// TIA Portal project "XSFW_TIA60401_A2" (V13)

(* hardware
DEVICE "SIMATIC 300(1)"  S7-300 station
   slot 0: "UR"  Rail  6ES7 390-1***0-0AA0
   slot 2: "CPU 315-2PN/DP"  CPU 315-2 PN/DP  6ES7 315-2EH14-0AB0  V3.1
      slot 2: "PN-IO"  PN-IO
         slot 1: "Puerto 1"  Port
         slot 2: "Puerto 2"  Port
   slot 4: "DI32xDC24V"  DI32xDC24V  6ES7 321-1BL00-0AA0
   slot 5: "DI32xDC24V_1"  DI32xDC24V  6ES7 321-1BL00-0AA0
   slot 6: "DI32xDC24V_2"  DI32xDC24V  6ES7 321-1BL00-0AA0
   slot 7: "DO32xDC24V/0.5A"  DO32xDC24V/0.5A  6ES7 322-1BL00-0AA0
   slot 8: "DO32xDC24V/0.5A_1"  DO32xDC24V/0.5A  6ES7 322-1BL00-0AA0
   slot 9: "AI8x13Bit"  AI8x13Bit  6ES7 331-1KF02-0AB0
   slot 10: "AI8x13Bit_1"  AI8x13Bit  6ES7 331-1KF02-0AB0
DEVICE "HMI-Chillers"  TP900 Comfort
   slot 0: "HMI"  HMI  6AV2 124-0JC01-0AX0  11.0.0
   slot 1: "HMI_RT_3"  TP900 Comfort  6AV2 124-0JC01-0AX0  11.0.0
   slot 5: "IE_CP_1"  PROFINET interface  IE_CP  V7.1.0
      slot 1: "PROFINET_Interfaz_1"  HMI IE SUBMODULE
         slot 1: "PORT_1"  HMI IE PORTMODULE 1  1.0.0.0
         slot 2: "PORT_2"  HMI IE PORTMODULE 1  1.0.0.0
   slot 7: "MPI/DP_CP_1"  HMI MPIDP  MPI-DP_CP  1.0.0.0
DEVICE "IM153-4PN"  S7-300 station
   slot 0: "UR"  Rail  6ES7 390-1***0-0AA0
   slot 0: "IM153-4PN"  IM 153-4PN  6ES7 153-4AA01-0XB0  V2.0
   slot 1: "DI32xDC24V"  DI32xDC24V  6ES7 321-1BL00-0AA0
   slot 2: "DI32xDC24V_2"  DI32xDC24V  6ES7 321-1BL00-0AA0
   slot 3: "DI32xDC24V_3"  DI32xDC24V  6ES7 321-1BL00-0AA0
   slot 4: "DO32xDC24V/0.5A_2"  DO32xDC24V/0.5A  6ES7 322-1BL00-0AA0
   slot 5: "DO32xDC24V/0.5A"  DO32xDC24V/0.5A  6ES7 322-1BL00-0AA0
   slot 6: "AI8x12Bit"  AI8 x 12 bits  6ES7 331-7KF02-0AB0
DEVICE "Cavaleto"  TP1200 Comfort
   slot 0: "HMI"  HMI  6AV2 124-0MC01-0AX0  13.0.1.0
   slot 1: "HMI_RT_1"  TP1200 Comfort  6AV2 124-0MC01-0AX0  13.0.1.0
   slot 5: "Cavaleto.IE_CP_1"  Interfaz PROFINET
      slot 1: "Interfaz PROFINET_1"  Interfaz PROFINET
         slot 1: "Port_1"  Port
         slot 2: "Port_2"  Port
   slot 7: "Cavaleto.MPI/DP_CP_1"  Interfaz MPI/DP
*)

// ===== PLC "CPU 315-2PN/DP"  CPU 315-2 PN/DP =====
// protected blocks, not shown: "FB_CTR_MOT", "FB_PRC_ALA", "FC_ANIM_MOTOR", "FC_CH_AI", "FC_MAQ_EST_16", "FC_PRC_ALA2", "FC_PRC_ALA3"

VAR_GLOBAL   // PLC tag table "Tabla de variables estándar"
   "Tag_1" AT %M7.0 : Bool;
   "Tag_2" AT %M7.1 : Bool;
   "Tag_3" AT %M7.2 : Bool;
   "Tag_4" AT %M7.3 : Bool;
   "Tag_5" AT %M7.4 : Bool;
   "Tag_6" AT %M500.0 : Bool;
   "Tag_7" AT %M900.0 : Bool;
   "Tag_9" AT %T15 : Timer;
   "Tag_10" AT %T16 : Timer;
   "Tag_11" AT %M55.0 : Bool;
   "Tag_12" AT %M330.3 : Bool;
   "Tag_13" AT %T80 : Timer;
   "flReqMch2" AT %M70.1 : Bool;
   "flReqMch3" AT %M70.2 : Bool;
   "flReqMch4" AT %M70.3 : Bool;
   "flReqMch5" AT %M70.4 : Bool;
   "Tag_18" AT %T62 : Timer;
   "Tag_19" AT %T61 : Timer;
   "Tag_20" AT %T60 : Timer;
   "Tag_21" AT %T70 : Timer;
   "Tag_22" AT %T71 : Timer;
   "Tag_23" AT %T72 : Timer;
   "Tag_24" AT %T73 : Timer;
   "Tag_25" AT %T74 : Timer;
   "Tag_26" AT %T24 : Timer;
   "Tag_27" AT %T10 : Timer;
   "Tag_28" AT %T11 : Timer;
   "Tag_29" AT %T12 : Timer;
   "Tag_30" AT %T13 : Timer;
   "Tag_31" AT %T14 : Timer;
   "Tag_32" AT %T26 : Timer;
   "Tag_33" AT %T28 : Timer;
   "Tag_34" AT %T30 : Timer;
   "Tag_35" AT %T32 : Timer;
   "Tag_36" AT %T34 : Timer;
   "Tag_37" AT %Q100.5 : Bool;
   "Tag_38" AT %M0.4 : Bool;
   "Tag_39" AT %Q104.4 : Bool;
   "Tag_40" AT %Q104.5 : Bool;
   "Tag_41" AT %Q101.1 : Bool;
   "Tag_42" AT %Q101.2 : Bool;
   "Tag_43" AT %Q101.3 : Bool;
   "Tag_44" AT %Q101.4 : Bool;
   "Tag_45" AT %Q101.5 : Bool;
   "Tag_46" AT %Q101.6 : Bool;
   "Tag_47" AT %Q101.7 : Bool;
   "Tag_48" AT %M25.0 : Bool;
   "Tag_49" AT %M25.1 : Bool;
   "Tag_50" AT %M25.2 : Bool;
   "Tag_51" AT %T35 : Timer;
   "Tag_52" AT %Q102.3 : Bool;
   "Tag_53" AT %Q102.4 : Bool;
   "Tag_54" AT %Q102.5 : Bool;
   "Tag_103" AT %M0.7 : Bool;
   "Tag_115" AT %M0.2 : Bool;
   "Tag_146" AT %M0.6 : Bool;
   "Tag_154" AT %M50.0 : Bool;
   "Tag_155" AT %M2.1 : Bool;
   "Tag_156" AT %M50.3 : Bool;
   "Tag_157" AT %M2.2 : Bool;
   "Tag_158" AT %M50.5 : Bool;
   "Tag_159" AT %M2.0 : Bool;
   "Tag_160" AT %Q69.1 : Bool;   // -
   "Tag_161" AT %M55.7 : Bool;
   "Tag_162" AT %M55.6 : Bool;
   "Latch_FT1" AT %M80.0 : Bool;   // Retención Flanco en Flujostato
   "Permiso_NO_FT1" AT %M80.1 : Bool;   // Permiso para trabajar sin FT1
   "Auxiliar_FT1" AT %M80.2 : Bool;
   "Auxiliar_Timer_FT1" AT %M80.3 : Bool;
   "Aviso 1" AT %M82.0 : Bool;
   "Aviso 2" AT %M82.1 : Bool;
   "Aviso 3" AT %M82.2 : Bool;
   "Aviso 4" AT %M82.3 : Bool;
   "Aviso 5" AT %M82.4 : Bool;
   "Aviso 13" AT %M82.6 : Bool;
   "Aviso 14" AT %M82.7 : Bool;
   "Aviso 23" AT %M83.0 : Bool;
   "Aviso 24" AT %M83.1 : Bool;
   "Aviso25" AT %M83.2 : Bool;
   "Aviso 26" AT %M83.3 : Bool;
   "Aviso 27" AT %M83.4 : Bool;
   "UltimoCmdMarcha" AT %M90.0 : Bool;
   "Tag_163" AT %T87 : Timer;
   "NotFirstScan" AT %M900.1 : Bool;
   "Tag_14" AT %M760.1 : Bool;
   "Tag_15" AT %M760.2 : Bool;
   "EnclavCompAltaConFlujostato" AT %M93.4 : Bool;
   "EstadoMantMC001" AT %MB761 : Byte;
   "EstadoMantMC002" AT %MB762 : Byte;
   "EstadoMantMC003" AT %MB763 : Byte;
   "EstadoMantMC004" AT %MB764 : Byte;
   "EstadoMantMC005" AT %MB765 : Byte;
   "EstadoMantMC006" AT %MB766 : Byte;
   "LimiteMantMC001_1" AT %M761.0 : Bool;
   "LimiteMantMC001_2" AT %M761.1 : Bool;
   "LimiteMantMC002_1" AT %M762.0 : Bool;
   "LimiteMantMC002_2" AT %M762.1 : Bool;
   "LimiteMantMC003_1" AT %M763.0 : Bool;
   "LimiteMantMC003_2" AT %M763.1 : Bool;
   "LimiteMantMC004_1" AT %M764.0 : Bool;
   "LimiteMantMC004_2" AT %M764.1 : Bool;
   "LimiteMantMC005_1" AT %M765.0 : Bool;
   "LimiteMantMC005_2" AT %M765.1 : Bool;
   "LimiteMantMC006_1" AT %M766.0 : Bool;
   "LimiteMantMC006_2" AT %M766.1 : Bool;
   "ProxMantMC001_1" AT %MD768 : DInt;
   "ProxMantMC002_1" AT %MD772 : DInt;
   "ProxMantMC003_1" AT %MD776 : DInt;
   "ProxMantMC004_1" AT %MD780 : DInt;
   "ProxMantMC005_1" AT %MD784 : DInt;
   "ProxMantMC006_1" AT %MD788 : DInt;
   "ProxMantMC001_2" AT %MD792 : DInt;
   "ProxMantMC002_2" AT %MD796 : DInt;
   "ProxMantMC003_2" AT %MD800 : DInt;
   "ProxMantMC004_2" AT %MD804 : DInt;
   "ProxMantMC005_2" AT %MD808 : DInt;
   "ProxMantMC006_2" AT %MD812 : DInt;
   "ProxMantMS050" AT %MD816 : DInt;
   "ProxMantMS051" AT %MD820 : DInt;
   "ProxMantMS052" AT %MD824 : DInt;
   "ProxMantMS053" AT %MD828 : DInt;
   "LimiteMantMS050" AT %M767.0 : Bool;
   "LimiteMantMS051" AT %M767.1 : Bool;
   "LimiteMantMS052" AT %M767.2 : Bool;
   "LimiteMantMS053" AT %M767.3 : Bool;
   "LimiteMantMS054_1" AT %M832.0 : Bool;
   "LimiteMantMS055_1" AT %M832.2 : Bool;
   "LimiteMantMS056_1" AT %M832.4 : Bool;
   "LimiteMantMS054_2" AT %M832.1 : Bool;
   "LimiteMantMS055_2" AT %M832.3 : Bool;
   "LimiteMantMS056_2" AT %M832.5 : Bool;
   "ProxMantMC060_1" AT %MD834 : DInt;
   "ProxMantMC061_1" AT %MD838 : DInt;
   "ProxMantMC062_1" AT %MD842 : DInt;
   "ProxMantMC063_1" AT %MD846 : DInt;
   "ProxMantMC064_1" AT %MD850 : DInt;
   "ProxMantMC065_1" AT %MD854 : DInt;
   "ProxMantMC060_2" AT %MD858 : DInt;
   "ProxMantMC061_2" AT %MD862 : DInt;
   "ProxMantMC062_2" AT %MD866 : DInt;
   "ProxMantMC063_2" AT %MD870 : DInt;
   "ProxMantMC064_2" AT %MD874 : DInt;
   "ProxMantMC065_2" AT %MD878 : DInt;
   "ProxMantMC060_3" AT %MD882 : DInt;
   "ProxMantMC061_3" AT %MD886 : DInt;
   "ProxMantMC062_3" AT %MD890 : DInt;
   "ProxMantMC063_3" AT %MD894 : DInt;
   "ProxMantMC064_3" AT %MD910 : DInt;
   "ProxMantMC065_3" AT %MD914 : DInt;
   "ProxMantMC060_4" AT %MD918 : DInt;
   "ProxMantMC061_4" AT %MD922 : DInt;
   "ProxMantMC062_4" AT %MD926 : DInt;
   "ProxMantMC063_4" AT %MD930 : DInt;
   "ProxMantMC064_4" AT %MD934 : DInt;
   "ProxMantMC065_4" AT %MD938 : DInt;
   "ProxMantMC060_5" AT %MD942 : DInt;
   "ProxMantMC061_5" AT %MD946 : DInt;
   "ProxMantMC062_5" AT %MD950 : DInt;
   "ProxMantMC063_5" AT %MD954 : DInt;
   "ProxMantMC064_5" AT %MD958 : DInt;
   "ProxMantMC065_5" AT %MD962 : DInt;
   "LimiteMantMC060_1" AT %M901.0 : Bool;
   "LimiteMantMC060_2" AT %M901.1 : Bool;
   "LimiteMantMC060_3" AT %M901.2 : Bool;
   "LimiteMantMC060_4" AT %M901.3 : Bool;
   "LimiteMantMC060_5" AT %M901.4 : Bool;
   "LimiteMantMC061_1" AT %M902.0 : Bool;
   "LimiteMantMC061_2" AT %M902.1 : Bool;
   "LimiteMantMC061_3" AT %M902.2 : Bool;
   "LimiteMantMC061_4" AT %M902.3 : Bool;
   "LimiteMantMC061_5" AT %M902.4 : Bool;
   "LimiteMantMC062_1" AT %M903.0 : Bool;
   "LimiteMantMC062_2" AT %M903.1 : Bool;
   "LimiteMantMC062_3" AT %M903.2 : Bool;
   "LimiteMantMC062_4" AT %M903.3 : Bool;
   "LimiteMantMC062_5" AT %M903.4 : Bool;
   "LimiteMantMC063_1" AT %M904.0 : Bool;
   "LimiteMantMC063_2" AT %M904.1 : Bool;
   "LimiteMantMC063_3" AT %M904.2 : Bool;
   "LimiteMantMC063_4" AT %M904.3 : Bool;
   "LimiteMantMC063_5" AT %M904.4 : Bool;
   "LimiteMantMC064_1" AT %M905.0 : Bool;
   "LimiteMantMC064_2" AT %M905.1 : Bool;
   "LimiteMantMC064_3" AT %M905.2 : Bool;
   "LimiteMantMC064_4" AT %M905.3 : Bool;
   "LimiteMantMC064_5" AT %M905.4 : Bool;
   "LimiteMantMC065_1" AT %M906.0 : Bool;
   "LimiteMantMC065_2" AT %M906.1 : Bool;
   "LimiteMantMC065_3" AT %M906.2 : Bool;
   "LimiteMantMC065_4" AT %M906.3 : Bool;
   "LimiteMantMC065_5" AT %M906.4 : Bool;
   "EstadoMantMC060" AT %MB901 : Byte;
   "EstadoMantMC061" AT %MB902 : Byte;
   "EstadoMantMC062" AT %MB903 : Byte;
   "EstadoMantMC063" AT %MB904 : Byte;
   "EstadoMantMC064" AT %MB905 : Byte;
   "ProxMantMS054_1" AT %MD966 : DInt;
   "ProxMantMS054_2" AT %MD970 : DInt;
   "ProxMantMS055_1" AT %MD974 : DInt;
   "ProxMantMS055_2" AT %MD978 : DInt;
   "EstadoMantSecBaja" AT %MB832 : Byte;
   "EnclavCompAltaPorTemp" AT %M93.5 : Bool;
   "FallTempCritEnclav" AT %M93.6 : Bool;
   "EntAnalCaudal" AT %IW266 : Word;
   "Tag_57" AT %MW982 : Word;
   "Tag_59" AT %MW984 : Word;
   "Tag_8" AT %M982.0 : Bool;
   "Tag_16" AT %M982.1 : Bool;
   "EntAnalPotencia" AT %IW264 : Word;
   "Tag_17" AT %T90 : Timer;
   "Tag_55" AT %T91 : Timer;
   "Tag_56" AT %M100.0 : Bool;
   "Tag_58" AT %M1000.0 : Bool;
   "Tag_60" AT %MW1010 : S5Time;
   "Tag_61" AT %MW1012 : S5Time;
   "MC003_EVP" AT %Q7.2 : Bool;   // Purga Bellis
   "Tag_63" AT %M1000.1 : Bool;
   "Tag_64" AT %T92 : Timer;
   "Tag_65" AT %T93 : Timer;
   "Tag_66" AT %MW1014 : S5Time;
   "Tag_67" AT %MW1016 : S5Time;
   "MC001_EVP" AT %Q7.3 : Bool;   // Purga ABC2
   "Tag_69" AT %M1000.2 : Bool;
   "Tag_70" AT %T94 : Timer;
   "Tag_71" AT %T95 : Timer;
   "Tag_72" AT %MW1018 : S5Time;
   "Tag_73" AT %MW1020 : S5Time;
   "MC002_EVP" AT %Q7.4 : Bool;   // Purga ABC3
   "Tag_75" AT %T96 : Timer;
   "Tag_76" AT %T97 : Timer;
   "MC004_EVP" AT %Q7.5 : Bool;   // Purga ABC4
   "Tag_78" AT %T98 : Timer;
   "Tag_79" AT %T99 : Timer;
   "MC005_EVP" AT %Q7.6 : Bool;   // Purga ABC5
   "Tag_62" AT %T100 : Timer;
   "MC006_EVP" AT %Q7.7 : Bool;   // Purga ABC1
   "Tag_68" AT %M1000.7 : Bool;
   "Tag_74" AT %T101 : Timer;
   "Tag_77" AT %T102 : Timer;
   "Tag_80" AT %T103 : Timer;
   "Tag_81" AT %T104 : Timer;
   "Tag_82" AT %T105 : Timer;
   "Tag_83" AT %T106 : Timer;
   "Tag_84" AT %T107 : Timer;
   "Tag_85" AT %I78.1 : Bool;
END_VAR

VAR_GLOBAL   // PLC tag table "STEP7 classic symbols"
   "MS055_MANT" AT %A4.1 : Bool;   // S BAJA SULLAIR 2-SEÑAL MODO MANTENIMIENTO / Secador 6 - SRD 1000 - Salida de Mantenimiento
   "MS055_Marcha" AT %A4.7 : Bool;   // S BAJA SULLAIR 2-CONTACTOR / Secador 6 - SRD 1000 - Salida de Marcha
   "MC006_TTB" AT %E2.2 : Bool;   // M COMPRESOR ALTA ABC1-TERMOSTATO AGUA / Secador 7 falla termico
   "MC006_TTA" AT %E2.3 : Bool;   // M COMPRESOR ALTA ABC1-TERMOSTATO AIRE / secador 8 falla termico
   "MT007-CO" AT %E66.0 : Bool;   // B SOPLADO L1-CONFIRMACIÓN DE MARCHA / Bomba Principal Chiller Soplado - Confirmación de Marcha
   "MT007-Marcha" AT %A66.0 : Bool;   // B SOPLADO L1-CONTACTOR / Accionamiento Bomba Intercambiador LINEA 1
   "MT007-TO" AT %E66.1 : Bool;   // B SOPLADO L1-TÉRMICO / Bomba Principal Chiller Soplado - Falla de Térmico
   "MT008-CO" AT %E66.2 : Bool;   // B SOPLADO L3 & MANOMEC-CONFIRMACIÓN DE MARCHA / Bomba Backup Chiller Soplado - Confirmación de Marcha
   "MT008-Marcha" AT %A66.1 : Bool;   // B SOPLADO L3 & MANOMEC-CONTACTOR / Accionamiento Bomba Intercambiador LINEA 2 Y MANOMEC
   "MT008-TO" AT %E66.3 : Bool;   // B SOPLADO L3 & MANOMEC-TÉRMICO / Bomba Backup Chiller Soplado - Falla de Térmico
   "MT009-CO" AT %E66.4 : Bool;   // B INT L3 Y L5-CONFIRMACIÓN DE MARCHA / Bomba Principal Chiller Envasado - Confirmación de Marcha
   "MT009-Marcha" AT %A66.2 : Bool;   // B INT L3 Y L5-CONTACTOR / Accionamiento Bomba Intercambiador LINEA 3 Y LINEA 5
   "MS052-TO" AT %E1.6 : Bool;   // M SECADOR ALTA ABC2-TÉRMICO / Secador 3-ABC 3- falla termico
   "MS052-VS1" AT %E9.4 : Bool;   // M SECADOR ALTA ABC2-PULSADOR PARADA / Secador 3 -ABC 3 - Falla de seguridades
   "MS052_MANT" AT %A3.6 : Bool;   // M SECADOR ALTA ABC2-SEÑAL MODO MANTENIMIENTO / Secador 2 - ABC 2 - Salida de Mantenimiento
   "FlancoMan2" AT %M322.7 : Bool;
   "FlancoMan3" AT %M323.0 : Bool;
   "FlancoMan4" AT %M323.1 : Bool;
   "FlancoMan5" AT %M323.2 : Bool;
   "FlancoManP1" AT %M323.3 : Bool;
   "FlancoManP2" AT %M323.4 : Bool;
   "FlancoManP3" AT %M323.5 : Bool;
   "FlancoManP4" AT %M323.6 : Bool;
   "FlancoManP5" AT %M323.7 : Bool;
   "TLUZ" AT %T17 : Timer;   // Tiempo Iluminación encendida
   "TOFF_SP1" AT %T44 : Timer;   // TOFF sopladora 1
   "TOFF_SP2" AT %T45 : Timer;   // TOFF Sopladora 2
   "TOFF_SP3" AT %T46 : Timer;   // TOFF Sopladora 3
   "TRetVCmp1" AT %T51 : Timer;   // Timer Retardo arranque de valvulas Compresor 1
   "TRetVCmp2" AT %T47 : Timer;   // Timer Retardo arranque de valvulas Compresor 2
   "TRetVCmp3" AT %T48 : Timer;   // Timer Retardo arranque de valvulas Compresor 3
   "TRetVCmp4" AT %T49 : Timer;   // Timer Retardo arranque de valvulas Compresor 4
   "TV1" AT %T53 : Timer;   // Timeout estando en vacío 1
   "TV2" AT %T36 : Timer;   // Timeout estando en vacío 2
   "TV3" AT %T37 : Timer;   // Timeout estando en vacío 3
   "TV4" AT %T38 : Timer;   // Timeout estando en vacío 4
   "FlaAux3" AT %M300.2 : Bool;   // Auxiliar arranque MC003
   "FlaAux4" AT %M300.3 : Bool;   // Auxiliar arranque MC004
   "FlaAux5" AT %M300.4 : Bool;   // Auxiliar arranque MC005
   "FlaAuxB1" AT %M300.5 : Bool;   // Auxiliar arranque MC061
   "FlaAuxB2" AT %M300.6 : Bool;   // Auxiliar arranque MC062
   "FlaAuxB3" AT %M300.7 : Bool;   // Auxiliar arranque MC063
   "FlaAuxB4" AT %M301.0 : Bool;   // Auxiliar arranque MC064
   "FlancoAuto1" AT %M324.0 : Bool;
   "FlancoAuto2" AT %M324.1 : Bool;
   "MP011-CO" AT %E67.2 : Bool;   // B BACKUP CH. SOPLADO-CONFIRMACIÓN DE MARCHA / Bomba Intercambiador LINEA 2 Y MANOMEC - Confirmación de Marcha
   "MP011-Marcha" AT %A66.5 : Bool;   // B BACKUP CH. SOPLADO-CONTACTOR / Accionamiento Bomba Backup Chiller Soplado
   "MP011-TO" AT %E67.3 : Bool;   // B BACKUP CH. SOPLADO-TÉRMICO / Bomba Intercambiador LINEA 2 Y MANOMEC - Falla de Térmico
   "MP012-CO" AT %E67.4 : Bool;   // B PRINC CH. ENVASADO-CONFIRMACIÓN DE MARCHA / Bomba Intercambiador LINEA 3 Y LINEA 5 - Confirmación de Marcha
   "MP012-Marcha" AT %A66.6 : Bool;   // B PRINC CH. ENVASADO-CONTACTOR / Accionamiento Bomba Principal Chiller Envasado
   "ArrMC061" AT %T81 : Timer;   // Timer arranque MC061
   "ArrMC062" AT %T82 : Timer;   // Timer arranque MC062
   "ArrMC063" AT %T83 : Timer;   // Timer arranque MC063
   "ArrMC064" AT %T84 : Timer;   // Timer arranque MC064
   "Arracando_MC002" AT %T27 : Timer;
   "Arrancando_MC001" AT %T25 : Timer;   // Delay para meter EV
   "Arrancando_MC004" AT %T31 : Timer;
   "Arrancando_MC005" AT %T33 : Timer;
   "Arrancando_mc003" AT %T29 : Timer;
   "BBA POZO" AT %A0.4 : Bool;   // BOMBA POZO- / BOMBA DE POZO
   "BMBTON2" AT %M69.3 : Bool;   // Bomba de torre 2 en funcionamiento
   "BMBTON2BMBTON" AT %M69.2 : Bool;   // Bomba de torre en funcionamiento
   "MC061-TO" AT %E11.5 : Bool;   // M COMPR BAJA SULLAIR 1-TÉRMICO / Compresor Baja SULL 1 - Falla de termico
   "MC005_ConfPurga" AT %E11.6 : Bool;   // ABC5 - Confirmación de electroválvula de purga. / Compresor Baja SULL 1 - Falla de seguridades
   "MC061_MANT" AT %A1.4 : Bool;   // M COMPR BAJA SULLAIR 1-SEÑAL MODO MANTENIMIENTO / Compresor Sullair1 Salida mantenimiento
   "MC061_MARCHA" AT %A1.5 : Bool;   // M COMPR BAJA SULLAIR 1-CONTACTOR / Comrpesor Sullair1 Salida de marcha
   "MC062-CO" AT %E10.3 : Bool;   // M COMPR BAJA SULLAIR 0-CONFIRMACIÓN DE MARCHA / Compresor Baja SULL 0- Conf. Marcha
   "MC062-TO" AT %E10.4 : Bool;   // M COMPR BAJA SULLAIR 0-TÉRMICO / Compresor Baja SULL 0- Falla de termico
   "MC062-VS1" AT %E10.5 : Bool;   // M COMPR BAJA SULLAIR 0-PULSADOR PARADA / Compresor Baja SULL 0- Falla de Seguridades
   "MC062_MANT" AT %A1.6 : Bool;   // M COMPR BAJA SULLAIR 0-SEÑAL MODO MANTENIMIENTO / Compresor XXX salida de mantenimiento
   "MC062_MARCHA" AT %A1.7 : Bool;   // M COMPR BAJA SULLAIR 0-CONTACTOR / Compresor XXX salida de marcha EX61
   "MC063-CO" AT %E10.6 : Bool;   // M COMPR BAJA ATLAS 3-CONFIRMACIÓN DE MARCHA / Compresor Baja ATLAS 3 - Conf.Marcha
   "MC063-TO" AT %E10.7 : Bool;   // M COMPR BAJA ATLAS 3-TÉRMICO / Compresor Baja ATLAS 3 - Falla de termico
   "IndicadorCmpAlta" AT %M310.4 : Bool;   // Indicador Aviso en Compresores de alta
   "IndicadorCmpBaja" AT %M310.2 : Bool;   // Indicador Aviso en Compresores de baja
   "IndicadorSecAlta" AT %M310.5 : Bool;   // Indicador Aviso en Secadores de alta
   "IndicadorSecBaja" AT %M310.3 : Bool;   // Indicador Aviso en Secadores de baja
   "IndicadorTorresCav" AT %M310.6 : Bool;   // Indicador Aviso en Torres cavalleto
   "IndicadorTorresCh" AT %M310.1 : Bool;   // Indicador Aviso en torres chillers
   "MC001" AT %A0.6 : Bool;   // M COMPRESOR ALTA ABC2-CONTACTOR / Compresor ABC2- Marcha-
   "MC001-CO" AT %E2.5 : Bool;   // M COMPRESOR ALTA ABC2-CONFIRMACIÓN DE MARCHA / Compresor ABC2-Confirmacion Marcha-
   "MC001-TO" AT %E2.6 : Bool;   // M COMPRESOR ALTA ABC2-TÉRMICO / Compresor ABC2-Falla Termico-
   "MC001_EV" AT %A2.0 : Bool;   // M COMPRESOR ALTA ABC2-ELECTROVÁLVULA / Electrovalvula libera carga MC001 (ABC2)
   "MC001_MANT" AT %A2.5 : Bool;   // M COMPRESOR ALTA ABC2-SEÑAL MODO MANTENIMIENTO / Compresor MC001 Salida Mantenimiento
   "MC002_ConfPurga" AT %E1.1 : Bool;   // ABC3 - Confirmación de electroválvula de purga. / Bomba de pozo -falla termico-
   "flReqMch1" AT %M70.0 : Bool;   // Flanco requerimiento de marcha compresor 1
   "TRetVCmp5" AT %T50 : Timer;   // Timer Retardo arranque de valvulas Compresor 5
   "FlancoTSinReq4" AT %M325.6 : Bool;
   "FlancoTSinReq5" AT %M325.7 : Bool;
   "FallaSensorTorresCH" AT %M77.7 : Bool;   // Falla en Sensor de Temperatura Torres de Chillers
   "FlaAux1" AT %M300.0 : Bool;   // Auxiliar arranque MC001
   "FlaAux2" AT %M300.1 : Bool;   // Auxiliar arranque MC002
   "Parada-MC062" AT %A6.0 : Bool;   // M COMPR BAJA SULLAIR 0-ORDEN PARADA / Parada MC062
   "Parada-MC063" AT %A5.7 : Bool;   // M COMPR BAJA ATLAS 3-ORDEN PARADA / Parada MC063
   "Parada-MC064" AT %A5.6 : Bool;   // M COMPR BAJA ATLAS 2-ORDEN PARADA / Parada MC064
   "P_PresALTA" AT %EW254 : Word;   // PresiónALTA
   "P_PresAlta2" AT %EW258 : Word;   // PresiónAlta2
   "P_PresBaja" AT %EW260 : Word;   // Presión Baja
   "Puls.Iluminati" AT %E7.5 : Bool;   // ILUMINACION-PULSADOR / Pulsador Iluminacion
   "Pulso0,5_Seg" AT %M1.0 : Bool;
   "Pulso100_Mseg" AT %M0.3 : Bool;
   "Pulso10_Seg" AT %M1.3 : Bool;
   "Pulso1_Seg" AT %M1.1 : Bool;
   "ErrCMQ1" AT %M320.5 : Bool;   // Error Concatenadoras Compresor 1
   "ErrCMQ2" AT %M320.6 : Bool;   // Error Concatenadoras Compresor 2
   "ErrCMQ3" AT %M320.7 : Bool;   // Error Concatenadoras Compresor 3
   "ErrCMQ4" AT %M321.0 : Bool;   // Error Concatenadoras Compresor 4
   "ErrCMQ5" AT %M321.1 : Bool;   // Error Concatenadoras Compresor 5
   "ErrCMQG" AT %M321.3 : Bool;   // Error Concatenadoras General
   "ErrPMQ1" AT %M320.0 : Bool;   // Error Prioritarias Compresor 1
   "ErrPMQ2" AT %M320.1 : Bool;   // Error Prioritarias Compresor 2
   "ErrPMQ3" AT %M320.2 : Bool;   // Error Prioritarias Compresor 3
   "ErrPMQ4" AT %M320.3 : Bool;   // Error Prioritarias Compresor 4
   "ErrPMQ5" AT %M320.4 : Bool;   // Error Prioritarias Compresor 5
   "BoosterAnimaMotor" AT %MB11 : Byte;   // Byte Animación Motor Booster
   "BoostMoManten" AT %M10.0 : Bool;   // Booster en modo Mantenimiento
   "BoostMoManual" AT %M10.1 : Bool;   // Booster en modo Manual
   "BoostMoAutoma" AT %M10.2 : Bool;   // Booster en modo Automático
   "BoosterAlarma" AT %M10.3 : Bool;   // Booster con Alarma Memorizada
   "BoostOrdMarch" AT %M10.4 : Bool;   // Booster con Orden de Marcha
   "BoostPlsManten" AT %M10.5 : Bool;   // Booster Pulsa Mantenimiento desde HMI
   "iConfMarBooster" AT %E3.7 : Bool;   // M BOOSTER 1-CONFIRMACIÓN DE MARCHA / Confirmaciónes Marcha serie motores Booster
   "iGMBooster" AT %E4.0 : Bool;   // M BOOSTER 1-GUARDAMOTOR / Confirmaciónes Guardamotores serie motores Booster
   "iPresostCtrl" AT %E7.6 : Bool;   // BOOSTERS (LOS DOS)-PRESOSTATO / Presostato de Control para Booster
   "iPresostPA" AT %E7.7 : Bool;   // BOOSTERS (LOS DOS)-PRESOSTATO PRESION ALTA / Presostato de "Presión Alta" para Booster
   "oMarBooster" AT %A7.0 : Bool;   // BOOSTER-CONTACTOR / Accionamiento Contactor Booster
   "FiltroPCtrlBooster" AT %T18 : Timer;   // Filtro de Presión de Control de Booster
   "FiltroPABooster" AT %T19 : Timer;   // Filtro de Presión Alta de Booster
   "Boost2OrdMarch" AT %M12.5 : Bool;   // Booster 2 con Orden de Marcha
   "Booster2Alarma" AT %M12.4 : Bool;   // Booster 2 con Alarma Memorizada
   "Boost2MoAutoma" AT %M12.3 : Bool;   // Booster 2 en modo Automático
   "Boost2MoManual" AT %M12.2 : Bool;   // Booster 2 en modo Manual
   "Boost2MoManten" AT %M12.1 : Bool;   // Booster 2 en modo Mantenimiento
   "BoostHabilit" AT %M12.0 : Bool;   // Habilitación Booster desde HMI
   "Boost2PlsManual" AT %M12.7 : Bool;   // Booster 2 Pulsa Manual desde HMI
   "Boost2PlsManten" AT %M12.6 : Bool;   // Booster 2 Pulsa Mantenimiento desde HMI
   "ReservaBooster_5" AT %M13.6 : Bool;
   "ReservaBooster_4" AT %M13.5 : Bool;
   "ReservaBooster_3" AT %M13.4 : Bool;
   "MS052_Marcha" AT %A4.4 : Bool;   // M SECADOR ALTA ABC2-CONTACTOR / Secador 3 - ABC 3 - Salida de Marcha
   "MS053-CO" AT %E4.4 : Bool;   // M SECADOR ALTA FARGON-CONFIRMACIÓN DE MARCHA / Secador 4 - Fargon -Conf.Marcha
   "MS053-TO" AT %E1.7 : Bool;   // M SECADOR ALTA FARGON-TÉRMICO / Secador 4-FARGON -falla termico
   "MS053-VS1" AT %E9.5 : Bool;   // M SECADOR ALTA FARGON-PULSADOR PARADA / Secador 4 -ABC Grande - Falla de seguridades
   "MS053_MANT" AT %A3.7 : Bool;   // M SECADOR ALTA FARGON-SEÑAL MODO MANTENIMIENTO / Secador 4- FARGON- Salida de Mantenimiento
   "MS053_Marcha" AT %A4.5 : Bool;   // M SECADOR ALTA FARGON-CONTACTOR / Secador 4 - FARGON - Salida de marcha
   "MS054-CO" AT %E4.5 : Bool;   // S BAJA SULLAIR 1-CONFIRMACIÓN DE MARCHA / Secador 5 -SRD850 - Conf.Marcha
   "MC006-CO" AT %E2.0 : Bool;   // M COMPRESOR ALTA ABC1-CONFIRMACIÓN DE MARCHA / Secador 5 - SRD 850 -falla termico
   "iConfMarBooster2" AT %E9.6 : Bool;   // M BOOSTER 2-CONFIRMACIÓN DE MARCHA / Confirmación de marcha Booster 2
   "MS054_MANT" AT %A4.0 : Bool;   // S BAJA SULLAIR 1-SEÑAL MODO MANTENIMIENTO / Secador 5 - SRD850 - Salida de Mantenimiento
   "MS054_Marcha" AT %A4.6 : Bool;   // S BAJA SULLAIR 1-CONTACTOR / Secador 5 - SRD850 - Salida de Marcha
   "MS055-CO" AT %E4.6 : Bool;   // S BAJA SULLAIR 2-CONFIRMACIÓN DE MARCHA / Secador 6 - SRD1000 - Conf.Marcha
   "MC006_PTB" AT %E2.1 : Bool;   // M COMPRESOR ALTA ABC1-PRESOSTATO AGUA / Secador 6 - SRD 1000-falla termico
   "Corneta" AT %A3.3 : Bool;   // -ALARMA / Bubuzella
   "MP019-CO" AT %E68.2 : Bool;   // BOMBA 2-CONFIRMACIÓN DE MARCHA / Bomba 2 Torres Enfriamiento - Confirmación de Marcha
   "MP019-Marcha" AT %A67.1 : Bool;   // BOMBA 2-CONTACTOR / Accionamiento Bomba 2 Torres Enfriamiento
   "MP019-TO" AT %E68.3 : Bool;   // BOMBA 2-TÉRMICO / Bomba 2 Torres Enfriamiento - Falla de Térmico
   "MP019_PA" AT %E8.3 : Bool;   // BOMBA 2-PULSADOR MARCHA / Bomba 2 Torre Cavalleto Pulsador Arranque
   "MP019_PP" AT %E8.4 : Bool;   // BOMBA 2-PULSADOR PARADA / Bomba 2 Torre Cavalleto Pulsador Parada
   "FlancoNoFal2" AT %M324.6 : Bool;
   "FlancoNoFal3" AT %M324.7 : Bool;
   "FlancoNoFal4" AT %M325.0 : Bool;
   "FlancoNoFal5" AT %M325.1 : Bool;
   "FlancoOsc1s" AT %M326.0 : Bool;
   "FlancoPSop1" AT %M326.4 : Bool;
   "FlancoPSop2" AT %M326.5 : Bool;
   "FlancoPSop3" AT %M326.6 : Bool;
   "FlancoTSinReq1" AT %M325.3 : Bool;
   "FlancoTSinReq2" AT %M325.4 : Bool;
   "FlancoTSinReq3" AT %M325.5 : Bool;
   "TV5" AT %T39 : Timer;   // Timeout estando en vacío 5
   "TdesefMC060" AT %T54 : Timer;   // Tiempo desconexión efectiva MC060
   "TdesefMC061" AT %T55 : Timer;   // Tiempo desconexión efectiva MC061
   "TdesefMC062" AT %T56 : Timer;   // Tiempo desconexión efectiva MC062
   "TdesefMC063" AT %T57 : Timer;   // Tiempo desconexión efectiva MC063
   "TdesefMC064" AT %T58 : Timer;   // Tiempo desconexión efectiva MC064
   "P_TemCav" AT %EW256 : Word;   // Temperatura Torres Cavaleto
   "TempTorresCH" AT %MD52 : Real;   // Temperatura Torres de Chillers Escalada
   "P_TempTorresCHILL" AT %EW286 : Word;   // Temperatura de agua torres de enfriamiento chillers
   "MC006_PTA" AT %E2.4 : Bool;   // M COMPRESOR ALTA ABC1-PRESOSTATO ACEITE / tomascorrientes falla termico
   "Torre_PE" AT %E9.1 : Bool;   // TORRE ENFR-PULS PARADA EMER / Pulsador de emergencia torre de enfriamiento
   "FlancoDEC5" AT %M322.5 : Bool;
   "FlancoINC1" AT %M321.4 : Bool;
   "FlancoINC2" AT %M321.5 : Bool;
   "FlancoINC3" AT %M321.6 : Bool;
   "FlancoINC4" AT %M321.7 : Bool;
   "FlancoINC5" AT %M322.0 : Bool;
   "FlancoMan1" AT %M322.6 : Bool;
   "ReservaBooster_2" AT %M13.3 : Bool;
   "ReservaBooster_1" AT %M13.2 : Bool;
   "Boost2Habilit" AT %M13.1 : Bool;   // Habilitación Booster 2 desde HMI
   "Boost2PlsAutoma" AT %M13.0 : Bool;   // Booster 2 Pulsa Automático desde HMI
   "oMarBooster2" AT %A7.1 : Bool;   // BOOSTER 2-CONTACTOR / Accionamiento Contactor Booster 2
   "ReservaBooster_6" AT %M13.7 : Bool;
   "Booster2AnimaMotor" AT %MB14 : Byte;   // Byte Animación Motor Booster 2
   "PrioridadBoost2" AT %MW334 : Int;   // Prioridad de Arranque Booster 2
   "PrioridadBoost1" AT %MW332 : Int;   // Prioridad de Arranque Booster 1
   "BoostAyuda" AT %M330.0 : Bool;   // Arrancar Booster de ayuda
   "BoostInvP" AT %M330.1 : Bool;   // Invertir Prioridad de Boosters
   "T_BoostHelp" AT %T21 : Timer;   // Tiempo para ayuda de Booster
   "T_OFFHelp" AT %T23 : Timer;   // Tiempo para quitar señal Ayuda Booster
   "FiltroPCtrlBooster2" AT %T22 : Timer;   // Filtro Control de Presión Booster 2
   "AuxTempBoos2" AT %MW338 : Int;   // Auxiliar para Temporización Horas Boost 2
   "AuxTempBoos1" AT %MW336 : Int;   // Auxiliar para Temporización Horas Boost 1
   "BoostPHor" AT %M330.2 : Bool;   // Control de Prioridades Boosters por Horas
   "P_iwPresBoosters" AT %EW262 : Word;   // Presión para el control de los Boosters
   "FallaUnBooster" AT %M330.4 : Bool;   // Falla en algún Booster
   "PresBoosters" AT %MD56 : Real;   // Presión Real para el control de los Boosters
   "BoostPrio2_ON" AT %M330.6 : Bool;   // Marcha Booster Prioridad 2
   "BoostPrio1_ON" AT %M330.5 : Bool;   // Marcha Booster Prioridad 1
   "BoostPrio2_OFF" AT %M331.0 : Bool;   // Parada Booster Prioridad 2
   "BoostPrio1_OFF" AT %M330.7 : Bool;   // Parada Booster Prioridad 1
   "CotaSupPresAna" AT %MD76 : Real;   // Cota Superior para lectura de Presión Analógica
   "ErrLectAna" AT %M331.1 : Bool;   // Error en Lectura analógica
   "MS050-CO" AT %E4.1 : Bool;   // M SECADOR ALTA ABC1-CONFIRMACIÓN DE MARCHA / Secador 1 -ABC Grande- Conf.Marcha
   "MS050-TO" AT %E1.4 : Bool;   // M SECADOR ALTA ABC1-TÉRMICO / Secador 1 - ABC Grande -falla termico
   "MS050-VS1" AT %E9.2 : Bool;   // M SECADOR ALTA ABC1-PULSADOR PARADA / Secador 1 - FARGON - Falla de Seguridades
   "MS050_MANT" AT %A3.4 : Bool;   // M SECADOR ALTA ABC1-SEÑAL MODO MANTENIMIENTO / Secador 1 - ABC Grande - Salida Mantenimiento
   "MS050_Marcha" AT %A4.2 : Bool;   // M SECADOR ALTA ABC1-CONTACTOR / Secador 1 - ABC Grande - Salida de Marcha
   "MS051-CO" AT %E4.2 : Bool;   // M SECADOR ALTA ABC3-CONFIRMACIÓN DE MARCHA / Secador 2 - ABC 2-Conf.Marcha
   "MS051-TO" AT %E1.5 : Bool;   // M SECADOR ALTA ABC3-TÉRMICO / Secador 2 - ABC2 -Falla termico
   "MS051-VS1" AT %E9.3 : Bool;   // M SECADOR ALTA ABC3-PULSADOR PARADA / Secador 2 -ABC 2 - Falla de Seguridades
   "MS051_MANT" AT %A3.5 : Bool;   // M SECADOR ALTA ABC3-SEÑAL MODO MANTENIMIENTO / Secador 2 - ABC 2 - Salida de Mantenimiento
   "MS051_Marcha" AT %A4.3 : Bool;   // M SECADOR ALTA ABC3-CONTACTOR / Secador 2 - ABC 2 - Salida de Marcha
   "MS052-CO" AT %E4.3 : Bool;   // M SECADOR ALTA ABC2-CONFIRMACIÓN DE MARCHA / Secador 3 - ABC-3 -Conf.Marcha
   "CHILL3-AL2" AT %E69.5 : Bool;   // CHILLER ENVASADO GRAND-ALARMA 2 / Chiller Envasado GRANDE - Alarma 2
   "CHILL3-MAX" AT %E69.7 : Bool;   // CHILLER ENVASADO GRAND-MAXIMA CAPACIDAD / Chiller Envasado GRANDE - Máxima Capacidad
   "CHILL3-RUN" AT %E69.6 : Bool;   // CHILLER ENVASADO GRAND- / Chiller Envasado GRANDE - En modo RUN
   "CHILL4-ACEITE" AT %E76.0 : Bool;   // CHILLER ENVASADO CHICO-FALLA ACEITE / Chiller Envasado CHICO - Alarma Aceite
   "CHILL4-RUN" AT %E76.3 : Bool;   // CHILLER ENVASADO CHICO- / Chiller Envasado CHICO - En Modo Funcionamiento
   "CHILL4-TEMP" AT %E76.1 : Bool;   // CHILLER ENVASADO CHICO-TEMPERATURA / Chiller Envasado CHICO - Alarma Temperatura
   "CHILL4-TERM1" AT %E76.2 : Bool;   // CHILLER ENVASADO CHICO-TÉRMICO / Chiller Envasado CHICO - Alarma Térmico
   "MP012-TO" AT %E67.5 : Bool;   // B PRINC CH. ENVASADO-TÉRMICO / Bomba Intercambiador LINEA 3 Y LINEA 5 - Falla de Térmico
   "MP013-CO" AT %E67.6 : Bool;   // B BACKUP CH. ENVASADO-CONFIRMACIÓN DE MARCHA / Bomba Intercambiador LINEA 1 Y MANOMEC - Confirmación de Marcha
   "MP013-Marcha" AT %A66.7 : Bool;   // B BACKUP CH. ENVASADO-CONTACTOR / Accionamiento Bomba Backup Chiller Envasado
   "MP013-TO" AT %E67.7 : Bool;   // B BACKUP CH. ENVASADO-TÉRMICO / Bomba Intercambiador LINEA 1 Y MANOMEC - Falla de Térmico
   "MP014" AT %A0.0 : Bool;   // BOMBA 1-CONTACTOR / BOMBA 1 TORRE -. marcha-
   "MP014-CO" AT %E0.0 : Bool;   // BOMBA 1-CONFIRMACIÓN DE MARCHA / BOMBA 1 TORRE ENF.-CONFIRMACION
   "FlancoAuto3" AT %M324.2 : Bool;
   "FlancoAuto4" AT %M324.3 : Bool;
   "FlancoAuto5" AT %M324.4 : Bool;
   "FlancoDEC1" AT %M322.1 : Bool;
   "FlancoDEC2" AT %M322.2 : Bool;
   "FlancoDEC3" AT %M322.3 : Bool;
   "FlancoDEC4" AT %M322.4 : Bool;
   "Pulso3_Seg" AT %M1.4 : Bool;
   "Pulso5_Seg" AT %M1.2 : Bool;
   "RetVLV1" AT %T63 : Timer;   // Retardo válvula 1
   "RetVLV2" AT %T64 : Timer;   // Retardo válvula 2
   "RetVLV3" AT %T65 : Timer;   // Retardo válvula 3
   "RetVLV3b" AT %T68 : Timer;   // Retardo válvula 3b
   "RetVLV4" AT %T66 : Timer;   // Retardo válvula 4
   "RetVLV5" AT %T67 : Timer;   // Retardo válvula 5
   "SirenaChillers" AT %A68.1 : Bool;   // CHILLER-CONTACTOR / SirenaChillers
   "T20" AT %T20 : Timer;   // Temporizador bloque de alarmas MTA
   "FT1_AGUA" AT %E8.0 : Bool;   // COMPRESORES-FUJOSTATO / Flujostato de Agua torre de enfriamiento cavalleto
   "Falla-FT1" AT %M20.0 : Bool;   // Falla Flujostato Agua Torre Cavalleto
   "MC063-VS1" AT %E11.0 : Bool;   // M COMPR BAJA ATLAS 3-PULSADOR PARADA / Compresor Baja ATLAS 3 - Falla de seguridades
   "MC063_MANT" AT %A5.0 : Bool;   // M COMPR BAJA ATLAS 3-SEÑAL MODO MANTENIMIENTO / Compresor ATLAS 3 salida de mantenimiento
   "MC063_MARCHA" AT %A5.1 : Bool;   // M COMPR BAJA ATLAS 3-CONTACTOR / Compresor ATLAS 3 salida de marcha
   "MC064-CO" AT %E11.1 : Bool;   // M COMPR BAJA ATLAS 2-CONFIRMACIÓN DE MARCHA / Compresor baja ATLAS 2- Conf.Marcha
   "MC064-TO" AT %E11.2 : Bool;   // M COMPR BAJA ATLAS 2-TÉRMICO / Compresor Baja ATLAS 2 - Falla de termico
   "A1.3" AT %A1.3 : Bool;   // - / Libre
   "AnulSir" AT %M600.0 : Bool;   // Anulación de Sirena Cavaleto
   "ArrMC001" AT %T75 : Timer;   // Timer arranque MC001
   "ArrMC002" AT %T76 : Timer;   // Timer arranque MC002
   "ArrMC003" AT %T77 : Timer;   // Timer arranque MC003
   "ArrMC004" AT %T78 : Timer;   // Timer arranque MC004
   "ArrMC005" AT %T79 : Timer;   // Timer arranque MC005
   "MC004_TTB" AT %E6.3 : Bool;   // M COMPRESOR ALTA ABC4-TERMOSTATO AGUA / Compresor ABC4 Alta Temperatura de agua
   "MC005" AT %A1.2 : Bool;   // M COMPRESOR ALTA ABC5-CONTACTOR / Compresor ABC5-. Marcha-(200 Kw)
   "MC005-CO" AT %E3.5 : Bool;   // M COMPRESOR ALTA ABC5-CONFIRMACIÓN DE MARCHA / Compresor ABC5-Confirmacion Marcha-(200 Kw)
   "MC005-TO" AT %E3.6 : Bool;   // M COMPRESOR ALTA ABC5-TÉRMICO / Compresor ABC5-Falla Termico--(200 Kw)
   "MC005_EV" AT %A2.4 : Bool;   // M COMPRESOR ALTA ABC5-ELECTROVÁLVULA / Electrovalvula libera carga MC005 (ABC5)